// TIA Portal project "Projeto caldeira - IHM" (V19)

(* hardware
DEVICE "S7-1200 station_2"  S7-1200 Station
   slot 0: "Rack_0"  S7-1200 Rack  Rack  V1.0
   slot 1: "PLC_2"  CPU 1215C DC/DC/DC  6ES7 215-1AG40-0XB0  V4.6
DEVICE "HMI_2"  KTP700 Basic PN
   slot 0: "HMI_2"  KTP700 Basic PN  6AV2 123-2GB03-0AX0  15.1.0.0
   slot 1: "HMI_RT_2"  KTP700 Basic PN  6AV2 123-2GB03-0AX0  15.1.0.0
   slot 5: "HMI_2.IE_CP_1"  PROFINET Interface  15.0.1.0
      slot 1: "PROFINET Interface_1"  PROFINET Interface
         slot 1: "Port_1"  Port
DEVICE "SCALANCE X005"  SCALANCE X-Station
   slot 0: "SCALANCE X rack"  Rail
   slot 0: "Switch_1"  6GK5 005-0BA00-1AB2  V1.0
*)

// ===== PLC "PLC_2"  CPU 1215C DC/DC/DC =====

VAR_GLOBAL   // PLC tag table "Dados"
   "Caldeira" AT %I0.0 : Bool;
   "Turbina_!" AT %I0.1 : Bool;
   "Turbina_2" AT %I0.2 : Bool;
   "Tanque_1" AT %I0.3 : Bool;
   "Tanque_2" AT %I0.4 : Bool;
END_VAR

DATA_BLOCK "Varáveis caldeira"   // DB1
{ S7_Optimized_Access := 'TRUE' }
VERSION : 0.1
   VAR
      Liga_caldeira : Bool;
      Liga_turbina : Bool;
      Liga_turbina_2 : Bool;
      Desliga_caldeira : Bool;
      Timer_1 : Bool;
      Timer_2 : Bool;
   END_VAR
BEGIN
END_DATA_BLOCK

DATA_BLOCK "Programação caldeira_DB"   // DB4
{ S7_Optimized_Access := 'TRUE' }
VERSION : 0.1
// stored: InstanceOfName Programação caldeira
"Programação caldeira"
BEGIN
END_DATA_BLOCK

// folder: System blocks/Program resources

DATA_BLOCK "timer 1"   // DB2
{ S7_Optimized_Access := 'TRUE' }
AUTHOR : Simatic
FAMILY : IEC
NAME : IEC_TMR
VERSION : 1.0
// stored: InstanceOfName IEC_TIMER
"IEC_TIMER"
BEGIN
END_DATA_BLOCK

DATA_BLOCK "IEC_Timer_0_DB"   // DB3
{ S7_Optimized_Access := 'TRUE' }
AUTHOR : Simatic
FAMILY : IEC
NAME : IEC_TMR
VERSION : 1.0
// stored: InstanceOfName IEC_TIMER
"IEC_TIMER"
BEGIN
END_DATA_BLOCK

// folder: (top level)

FUNCTION_BLOCK "Programação caldeira"   // FB1, LAD
{ S7_Optimized_Access := 'TRUE' }
VERSION : 0.1
BEGIN

REGION Network 1
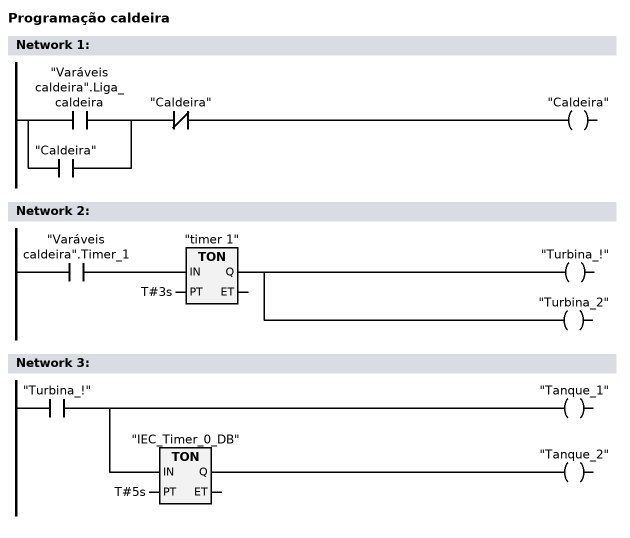
   RUNG wire#powerrail
      Contact( "Varáveis caldeira".Liga_caldeira )
      wire#w1
      I_Contact( "Caldeira" )
      Coil( "Caldeira" )
   END_RUNG
   RUNG wire#powerrail
      Contact( "Caldeira" )
   END_RUNG wire#w1
   // the same network as SCL:
   "Caldeira" := ("Varáveis caldeira".Liga_caldeira OR "Caldeira") AND NOT "Caldeira";
END_REGION

REGION Network 2
   "timer 1".TON(IN := "Varáveis caldeira".Timer_1, PT := T#3s);
   "Turbina_!" := "timer 1".Q;
   "Turbina_2" := "timer 1".Q;
END_REGION

REGION Network 3
   "Tanque_1" := "Turbina_!";
   "IEC_Timer_0_DB".TON(IN := "Turbina_!", PT := T#5s);
   "Tanque_2" := "IEC_Timer_0_DB".Q;
END_REGION
END_FUNCTION_BLOCK

ORGANIZATION_BLOCK "Main"   // OB1, LAD, ProgramCycle
TITLE = "Main Program Sweep (Cycle)"
{ S7_Optimized_Access := 'TRUE' }
VERSION : 0.1
   VAR_INPUT
      Initial_Call : Bool;   // Initial call of this OB
      Remanence : Bool;   // =True, if remanent data are available
   END_VAR
BEGIN

REGION Network 1
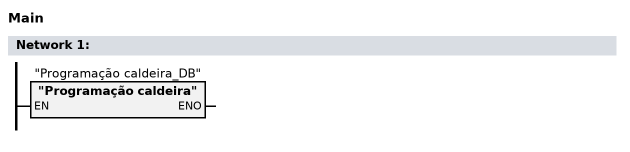
   RUNG wire#powerrail
      "Programação caldeira_DB"()
   END_RUNG
   // the same network as SCL:
   "Programação caldeira_DB"();   // "Programação caldeira"
END_REGION
END_ORGANIZATION_BLOCK

(* ===== HMI "HMI_RT_2" =====
system functions are stored by id; their names below are inferred from use
connection "HMI_Connection_2": ETHERNET, SMART_S7_1200_OMS

HMI tags "Default tag table"
   "Tag_ScreenNumber" : UInt, internal
   "Varáveis caldeira_Liga_caldeira" : Bool = PLC "Varáveis caldeira".Liga_caldeira, 1 s
   "Turbina_!" : Bool = PLC Turbina_! AT %I0.1, 1 s
   "Turbina_2" : Bool = PLC Turbina_2 AT %I0.2, 1 s
   "Tanque_1" : Bool = PLC Tanque_1 AT %I0.3, 1 s
   "Tanque_2" : Bool = PLC Tanque_2 AT %I0.4, 1 s

Template "Template_1" 800x480
   Button "Exit" at 714,429 size 71x50; TextOff 'Exit'; PictureOff "ExitRuntime_KTP700_Basic_PN_TR"; PictureOn "ExitRuntime_KTP700_Basic_PN_TR"
      on Release: StopRuntime(0)
   Button "Template_Button" at 614,429 size 71x50; TextOff 'Text'
   Button "Template_Button_1" at 514,429 size 71x50; TextOff 'Text'
   Button "Template_Button_2" at 414,429 size 71x50; TextOff 'Text'
   Button "Template_Button_3" at 314,429 size 71x50; TextOff 'Text'
   Button "Template_Button_4" at 214,429 size 71x50; TextOff 'Text'
   Button "Template_Button_5" at 114,429 size 71x50; TextOff 'Text'
   Button "Start screen" at 14,429 size 71x50; TextOff 'Start screen'; PictureOff "NavigateHome_KTP700_Basic_PN_TR"; PictureOn "NavigateHome_KTP700_Basic_PN_TR"
      on Release: ActivateScreen("Root screen", 0)
   SymbolicIOField "Symbolic_IO_Field_Screen" at 93,9 size 600x33; TextOff '0'; TextOn '1'; TextList "TextList_ScreenNames"
      ProcessValue <- "Tag_ScreenNumber"
      on Change: ActivateScreenByNumber("Tag_ScreenNumber", 0)
   DateTimeField "HmiScreenItemData" at 695,25 size 105x25
   DateTimeField "HmiScreenItemData_1" at 695,0 size 105x25
   GraphicView "Logo" at 0,0 size 91x51; Picture "Logo of HMI_2"

screen "Root screen" 800x480, template "Template_1"
   on GenerateScreen: SetTag("Tag_ScreenNumber", 1)
   TextField "HmiScreenItemData" at 80,225 size 640x25; Text 'Welcome to HMI_2 (KTP700 Basic+ PN)!'

screen "Principal" 800x480
   TextField "Text field_1" at 259,20 size 258x39; Text 'Controle Caldeira'
   Button "Button_1" at 295,162 size 187x62; TextOff 'Liga'
      on Click: SetBit("Varáveis caldeira_Liga_caldeira")
   Circle "Circle_3" at 236,357 size 48x48
      Appearance <- "Turbina_2"
   Circle "Circle_4" at 172,357 size 48x48
      Appearance <- "Turbina_!"
   TextField "Text field_2" at 184,320 size 88x27; Text 'Turbinas'
   TextField "Text field_3" at 188,368 size 15x23; Text '1'
   TextField "Text field_4" at 252,369 size 15x23; Text '2'
   Rectangle "Rectangle_2" at 293,231 size 192x9
      Appearance <- "Varáveis caldeira_Liga_caldeira"
   TextField "Text field_5" at 359,321 size 75x27; Text 'Válvula'
   Circle "Circle_1" at 517,355 size 48x48
      Appearance <- "Tanque_1"
   Circle "Circle_5" at 585,355 size 48x48
      Appearance <- "Tanque_2"
   TextField "Text field_6" at 536,323 size 75x27; Text 'Tanque'
   TextField "Text field_7" at 533,366 size 15x23; Text '1'
   TextField "Text field_8" at 601,367 size 15x23; Text '2'
*)